// TIA Portal project "Lagerregal_6" (V20)

(* hardware
DEVICE "S7-1500/ET200MP-Station_1"  S7-1500 station
   slot 0: "Profilschiene_0"  Rack  6ES7 590-1***0-0AA0
   slot 1: "PLC_1"  CPU 1513-1 PN  6ES7 513-1AM03-0AB0  V4.0
      slot 3: "CPU-Display_1"  6ES7591-1AA00-0AA0
      slot 32768: "PROFINET-Schnittstelle_1"  X1
         slot 32769: "Port_1"  X1 P1
         slot 32770: "Port_2"  X1 P2
      slot 34817: "Virtual CP interface port_1"  Virtual CP interface port  Virtual CP interface port FW V4.0
   slot 2: "DI 16x24VDC BA_1"  DI 16x24VDC BA  6ES7 521-1BH10-0AA0  V1.1
   slot 3: "DQ 16x24VDC/0.5A ST_1"  DQ 16x24VDC/0.5A ST  6ES7 522-1BH00-0AB0  V2.0
   slot 4: "AI 8xU/I/R/RTD BA_2"  AI 8xU/I/R/RTD BA  6ES7 531-7QF00-0AB0  V1.0
   slot 5: "AI 8xU/I/R/RTD BA_1"  AI 8xU/I/R/RTD BA  6ES7 531-7QF00-0AB0  V1.0
DEVICE "HMI_1"  TP700 Comfort
   slot 0: "HMI_1"  TP700 Comfort  6AV2 124-0GC01-0AX0  17.0.0.0
   slot 1: "HMI_RT_1"  TP700 Comfort  6AV2 124-0GC01-0AX0  17.0.0.0
   slot 5: "HMI_1.IE_CP_1"  PROFINET Interface  17.0.0.0
      slot 1: "PROFINET Schnittstelle_1"  PROFINET Interface
         slot 1: "Port_1"  Port
         slot 2: "Port_2"  Port
   slot 7: "HMI_1.MPI/DP_CP_1"  MPI/DP Interface  17.0.0.0
*)

// ===== PLC "PLC_1"  CPU 1513-1 PN =====

VAR_GLOBAL   // PLC tag table "Standard-Variablentabelle"
   "Clock_Byte" AT %MB0 : Byte;
   "Clock_10Hz" AT %M0.0 : Bool;
   "Clock_5Hz" AT %M0.1 : Bool;
   "Clock_2.5Hz" AT %M0.2 : Bool;
   "Clock_2Hz" AT %M0.3 : Bool;
   "Clock_1.25Hz" AT %M0.4 : Bool;
   "Clock_1Hz" AT %M0.5 : Bool;
   "Clock_0.625Hz" AT %M0.6 : Bool;
   "Clock_0.5Hz" AT %M0.7 : Bool;
END_VAR

VAR_GLOBAL CONSTANT   // PLC tag table "Standard-Variablentabelle"
   "Fachhoehe" : Int := 4800;
   "Fachbreite" : Int := 2962;
   "Offset-Z" : Int := 1800;
   "Offset-X" : Int := 3952;
   "Faecher_pro_Zeile" : Int := 9;
   "Faecher_pro_Spalte" : Int := 6;
   "Anheben_Absenken" : Int := 1000;
END_VAR

VAR_GLOBAL   // PLC tag table "Eingaenge"
   "S1" AT %I0.0 : Bool;   // Not-Aus
   "S2" AT %I0.1 : Bool;   // Anlage ein
   "S3" AT %I0.2 : Bool;   // Starttaster
   "1B1" AT %I0.3 : Bool;   // Sensor 1. Einlassband Anfang
   "1B2" AT %I0.4 : Bool;   // Sensor 1. Einlassband Ende
   "2B1" AT %I0.5 : Bool;   // Sensor 2. Einlassband Anfang
   "2B2" AT %I0.6 : Bool;   // Sensor 2. Einlassband Ende
   "3B1" AT %I0.7 : Bool;   // Sensor 3. Einlassband
   "4B1" AT %I1.0 : Bool;   // Sensor 1. Auslassband
   "5B1" AT %I1.1 : Bool;   // Sensor 2. Auslassband
   "6B1" AT %I1.2 : Bool;   // Endlage Gabel-Kran 1 (links)
   "6B2" AT %I1.3 : Bool;   // Endlage Gabel-Kran 1 (rechts)
   "6B3" AT %I1.4 : Bool;   // Endlage Gabel-Kran 1 (mitte)
   "7B1" AT %I1.5 : Bool;   // Endlage Gabel-Kran 2 (links)
   "7B2" AT %I1.6 : Bool;   // Endlage Gabel-Kran 2 (rechts)
   "7B3" AT %I1.7 : Bool;   // Endlage Gabel-Kran 2 (mitte)
   "2B3" AT %EW30 : Int;   // Kamera am Einlass (Bauteilerkennung)
   "6B4" AT %EW32 : Int;   // X-Achse Kran 1 Ist-Pos
   "6B5" AT %EW34 : Int;   // Z-Achse Kran 1 Ist-Pos
   "7B4" AT %EW36 : Int;   // X-Achse Kran 2 Ist-Pos
   "7B5" AT %EW38 : Int;   // Z-Achse Kran 2 Ist-Pos
END_VAR

VAR_GLOBAL   // PLC tag table "Ausgaenge"
   "H3" AT %Q0.2 : Bool;   // Starttasterleuchte
   "1M1" AT %Q0.3 : Bool;   // 1. Einlassband
   "2M1" AT %Q0.5 : Bool;   // 2. Einlassband
   "3M1" AT %Q0.7 : Bool;   // 3. Einlassband
   "4M1" AT %Q1.0 : Bool;   // 1. Auslassband
   "5M1" AT %Q1.1 : Bool;   // 2. Auslassband
   "6M1" AT %Q1.2 : Bool;   // Gabel-Kran 1 (links)
   "6M2" AT %Q1.3 : Bool;   // Gabel-Kran 1 (rechts)
   "7M1" AT %Q1.5 : Bool;   // Gabel-Kran 2 (links)
   "7M2" AT %Q1.6 : Bool;   // Gabel-Kran 2 (rechts)
   "6M4" AT %AW32 : Int;   // X-Achse Kran 1 Soll-Pos
   "6M5" AT %AW34 : Int;   // Z-Achse Kran 1 Soll-Pos
   "7M4" AT %AW36 : Int;   // X-Achse Kran 2 Soll-Pos
   "7M5" AT %AW38 : Int;   // Z-Achse Kran 2 Soll-Pos
END_VAR

TYPE "typKran_Pos"
   STRUCT
      "X-Ist" : Int;   // X-Achse Kran Ist-Pos
      "X-Soll" : Int;   // X-Achse Kran Soll-Pos
      "X-Rechnen" : Int;   // Zwischenvariable um neue X-Achsen Soll-Pos zu bestimmen
      "X-Skaliert" : Real;
      "Z-Ist" : Int;   // Z-Achse Kran Ist-Pos
      "Z-Soll" : Int;   // Z-Achse Kran Soll-Pos
      "Z-Rechnen" : Int;   // Zwischenvariable um neue Z-Achsen Soll-Pos zu bestimmen
      "Z-Skaliert" : Real;
   END_STRUCT;
END_TYPE

TYPE "typLagerplatz"
   STRUCT
      Flags : Struct
         Belegt : Bool;
         In_Benutzung : Bool;
      END_STRUCT;
      Artikel_Nr : Int;
      Bauteil : Int;
      Zeitstempel : DTL;
      MHD : Date;
   END_STRUCT;
END_TYPE

TYPE "typSchritte"
   STRUCT
      Schritt_Init : Bool;
      Kran : Struct
         Schritt_1 : Bool;
         Schritt_2 : Bool;
         Schritt_3 : Bool;
         Schritt_4 : Bool;
         Schritt_5 : Bool;
      END_STRUCT;
      Kran_Beladen : Struct
         Schritt_1 : Bool;
         Schritt_2 : Bool;
         Schritt_3 : Bool;
         Schritt_4 : Bool;
      END_STRUCT;
      Kran_Entladen : Struct
         Schritt_1 : Bool;
         Schritt_2 : Bool;
         Schritt_3 : Bool;
         Schritt_4 : Bool;
      END_STRUCT;
   END_STRUCT;
END_TYPE

DATA_BLOCK "HMI_Schnittstelle"   // DB100
{ S7_Optimized_Access := 'TRUE' }
VERSION : 0.1
   VAR
      Eingaenge : Struct
         S1 : Bool;   // Not-Aus
         S2 : Bool;   // Anlage ein
         S3 : Bool;   // Starttaster
         "1B1" : Bool;   // Sensor 1. Einlassband Anfang
         "1B2" : Bool;   // Sensor 1. Einlassband Ende
         "2B1" : Bool;   // Sensor 2. Einlassband Anfang
         "2B2" : Bool;   // Sensor 2. Einlassband Ende
         "2B3" : Int;
         "3B1" : Bool;   // Sensor 3. Einlassband
         "4B1" : Bool;   // Sensor 1. Auslassband
         "5B1" : Bool;   // Sensor 2. Auslassband
         "6B1" : Bool;   // Endlage Gabel-Kran 1 (links)
         "6B2" : Bool;   // Endlage Gabel-Kran 1 (rechts)
         "6B3" : Bool;   // Endlage Gabel-Kran 1 (mitte)
         "7B1" : Bool;   // Endlage Gabel-Kran 2 (links)
         "7B2" : Bool;   // Endlage Gabel-Kran 2 (rechts)
         "7B3" : Bool;   // Endlage Gabel-Kran 2 (mitte)
      END_STRUCT;
      Ausgaenge : Struct
         H1 : Bool;   // Starttasterleuchte
         "1M1" : Bool;   // 1. Einlassband
         "2M1" : Bool;   // 2. Einlassband
         "3M1" : Bool;   // 3. Einlassband
         "4M1" : Bool;   // 1. Auslassband
         "5M1" : Bool;   // 2. Auslassband
         "6M1" : Bool;   // Gabel-Kran 1 (links)
         "6M2" : Bool;   // Gabel-Kran 1 (rechts)
         "7M1" : Bool;   // Gabel-Kran 2 (links)
         "7M2" : Bool;   // Gabel-Kran 2 (rechts)
      END_STRUCT;
      Betriebsart : Struct
         Hand : Bool;
         Automatik : Bool;
         Stopp : Bool;
         Einrichten : Bool;
      END_STRUCT;
      Anlagendaten : Struct
         Schrittnummer : UInt;
         Fach_ansteuern : Bool;
         Fach : Int := 1;
         Bauteil : Int;
         Regalplatz_frei : Bool;
         Band_ein : Array[1..3] of Int;
         Band_aus : Array[1..2] of Int;
      END_STRUCT;
      Kraene : Struct
         Kran_1 : Struct
            Kran_Pos : "typKran_Pos";
            Kran_Schritt_Nr : Int;
            Schritt_Beladen : Int;
            Schritt_Entladen : Int;
            Grundstellung : Bool;
            Heimposition : Bool;
            Steht : Bool;
            Beladen : Bool;
         END_STRUCT;
         Kran_2 : Struct
            Kran_Pos : "typKran_Pos";
            Kran_Schritt_Nr : Int;
            Schritt_Beladen : Int;
            Schritt_Entladen : Int;
            Grundstellung : Bool;
            Heimposition : Bool;
            Steht : Bool;
            Beladen : Bool;
         END_STRUCT;
      END_STRUCT;
      HMI : Struct
         "X-Pos" : Bool;   // X-Achse-Inkrement erhöhen Schalter
         "X-Neg" : Bool;   // X-Achse-Inkrement verringern Schalter
         "Z-Pos" : Bool;   // Z-Achse-Inkrement erhöhen Schalter
         "Z-Neg" : Bool;   // Z-Achse-Inkrement verringern Schalter
         Inkrement : UInt;   // Inkrement Schrittgröße für Achsen
      END_STRUCT;
      Bitmeldungen : Word;
   END_VAR
BEGIN
   // Kraene.Kran_1.Kran_Pos."X-Ist" : X-Achse Kran 1 Ist-Pos
   // Kraene.Kran_1.Kran_Pos."Z-Ist" : Z-Achse Kran 1 Ist-Pos
   // Kraene.Kran_2.Kran_Pos."X-Ist" : X-Achse Kran 2 Ist-Pos
   // Kraene.Kran_2.Kran_Pos."Z-Ist" : Z-Achse Kran 2 Ist-Pos
   // Kraene.Kran_1.Kran_Pos."X-Soll" : X-Achse Kran 1 Soll-Pos
   // Kraene.Kran_1.Kran_Pos."Z-Soll" : Z-Achse Kran 1 Soll-Pos
   // Kraene.Kran_2.Kran_Pos."X-Soll" : X-Achse Kran 2 Soll-Pos
   // Kraene.Kran_2.Kran_Pos."Z-Soll" : Z-Achse Kran 2 Soll-Pos
END_DATA_BLOCK

DATA_BLOCK "Warenlager"   // DB101
{ S7_Optimized_Access := 'TRUE' }
VERSION : 0.1
   VAR
      Lager : Array[0..54] of "typLagerplatz";
   END_VAR
BEGIN
END_DATA_BLOCK

// folder: Anlagedaten

DATA_BLOCK "IDB_Anlage"   // DB1
{ S7_Optimized_Access := 'TRUE' }
VERSION : 0.1
// stored: InstanceOfName Ein_Anlage
"Ein_Anlage"
BEGIN
END_DATA_BLOCK

// folder: Bandsteuerung

DATA_BLOCK "IDB_Baender"   // DB20
{ S7_Optimized_Access := 'TRUE' }
VERSION : 0.1
// stored: InstanceOfName Ein_Baender
"Ein_Baender"
BEGIN
END_DATA_BLOCK

DATA_BLOCK "IDB_Bandsteuerung"   // DB21
{ S7_Optimized_Access := 'TRUE' }
VERSION : 0.1
// stored: InstanceOfName Bandsteuerung
"Bandsteuerung"
BEGIN
END_DATA_BLOCK

// folder: HMI

DATA_BLOCK "IDB_Einrichtbetrieb"   // DB3
{ S7_Optimized_Access := 'TRUE' }
VERSION : 0.1
// stored: InstanceOfName Prog_Einrichtbetrieb
"Prog_Einrichtbetrieb"
BEGIN
END_DATA_BLOCK

DATA_BLOCK "IDB_HMI"   // DB10
{ S7_Optimized_Access := 'TRUE' }
VERSION : 0.1
// stored: InstanceOfName Ein_HMI
"Ein_HMI"
BEGIN
END_DATA_BLOCK

// folder: Kransteuerung

DATA_BLOCK "IDB_Kran_beladen"   // DB25
{ S7_Optimized_Access := 'TRUE' }
VERSION : 0.1
// stored: InstanceOfName FC_Kran_beladen
"FC_Kran_beladen"
BEGIN
END_DATA_BLOCK

DATA_BLOCK "IDB_Kran"   // DB30
{ S7_Optimized_Access := 'TRUE' }
VERSION : 0.1
// stored: InstanceOfName Ein_Kran
"Ein_Kran"
BEGIN
END_DATA_BLOCK

DATA_BLOCK "IDB_Automatik_einlagern"   // DB50
{ S7_Optimized_Access := 'TRUE' }
VERSION : 0.1
// stored: InstanceOfName Prog_Automatik_einlagern
"Prog_Automatik_einlagern"
BEGIN
END_DATA_BLOCK

DATA_BLOCK "IDB_Automatik_auslagern"   // DB60
{ S7_Optimized_Access := 'TRUE' }
VERSION : 0.1
// stored: InstanceOfName Prog_Automatik_auslagern
"Prog_Automatik_auslagern"
BEGIN
END_DATA_BLOCK

// folder: (top level)

FUNCTION_BLOCK "Prog_Schrittkette"   // FB1234, FBD
{ S7_Optimized_Access := 'TRUE' }
VERSION : 0.1
   VAR_INPUT
      eAutomatik : Bool;   // Automatikmodus
      eAusschalten : Bool;   // Ausschalten der Schrittkette
      T_1_2 : Bool;
      T_2_3 : Bool;
      T_3_4 : Bool := TRUE;
      T_4_5 : Bool := TRUE;
      T_5_6 : Bool := TRUE;
      T_6_7 : Bool := TRUE;
      T_7_8 : Bool := TRUE;
      T_8_9 : Bool := TRUE;
      T_9_10 : Bool := TRUE;
      T_10_1 : Bool := TRUE;
   END_VAR
   VAR_OUTPUT
      aSchrittnummer : Int;
   END_VAR
   VAR
      Step_1 : Bool;
      Step_2 : Bool;
      Step_3 : Bool;
      Step_4 : Bool;
      Step_5 : Bool;
      Step_6 : Bool;
      Step_7 : Bool;
      Step_8 : Bool;
      Step_9 : Bool;
      Step_10 : Bool;
   END_VAR
BEGIN

REGION Network 1: Step 1
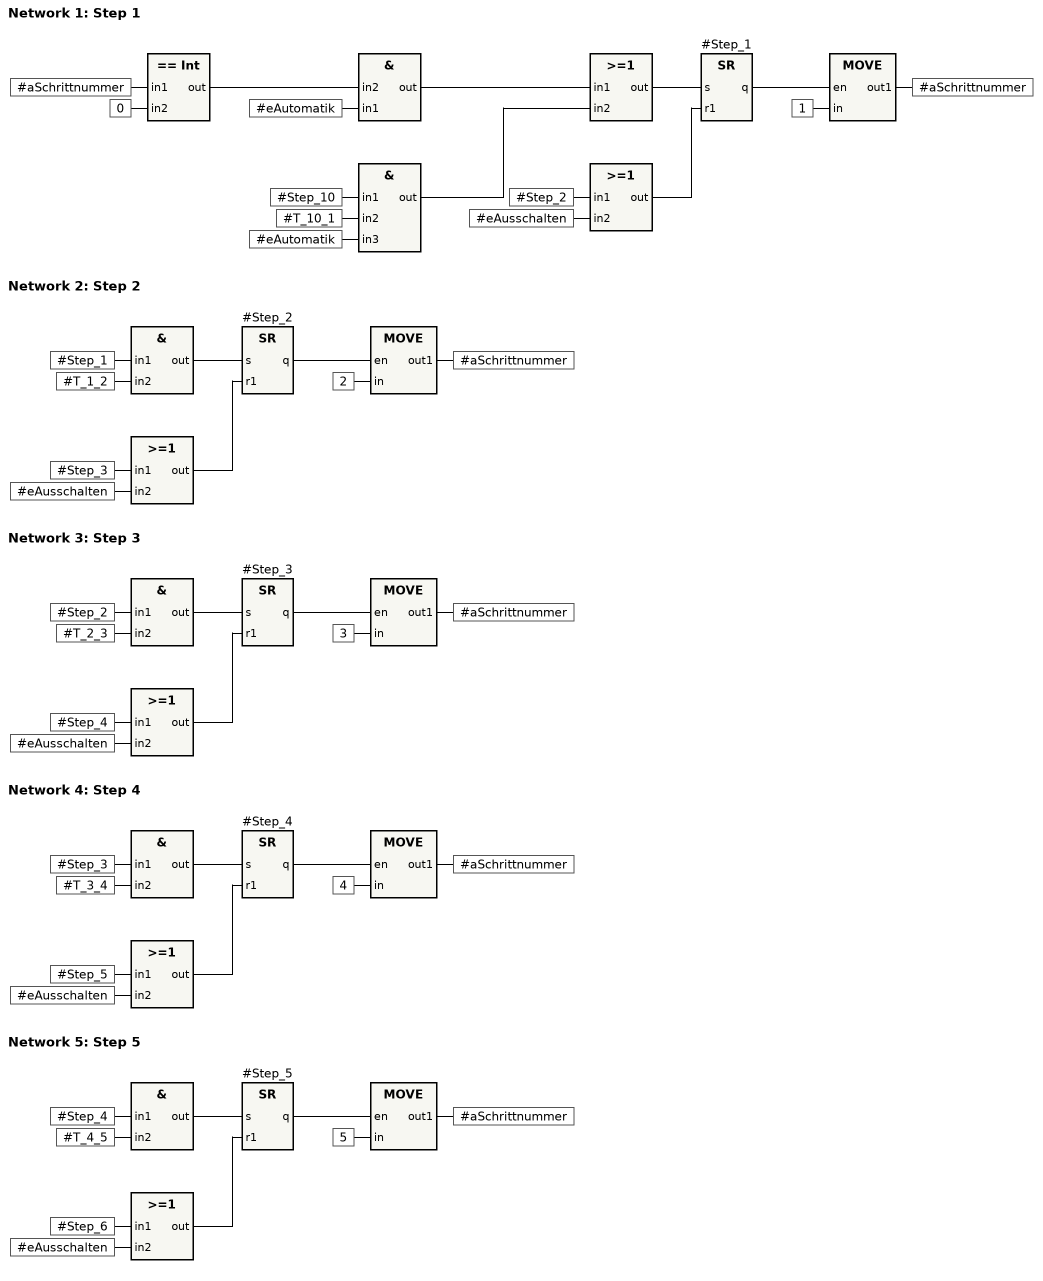
   IF ((#aSchrittnummer = 0) AND #eAutomatik) OR (#Step_10 AND #T_10_1 AND #eAutomatik) THEN
       #Step_1 := TRUE;   // SR flip-flop
   END_IF;
   IF #Step_2 OR #eAusschalten THEN #Step_1 := FALSE; END_IF;
   IF #Step_1 THEN #aSchrittnummer := 1; END_IF;
END_REGION

REGION Network 2: Step 2
   IF #Step_1 AND #T_1_2 THEN
       #Step_2 := TRUE;   // SR flip-flop
   END_IF;
   IF #Step_3 OR #eAusschalten THEN #Step_2 := FALSE; END_IF;
   IF #Step_2 THEN #aSchrittnummer := 2; END_IF;
END_REGION

REGION Network 3: Step 3
   IF #Step_2 AND #T_2_3 THEN
       #Step_3 := TRUE;   // SR flip-flop
   END_IF;
   IF #Step_4 OR #eAusschalten THEN #Step_3 := FALSE; END_IF;
   IF #Step_3 THEN #aSchrittnummer := 3; END_IF;
END_REGION

REGION Network 4: Step 4
   IF #Step_3 AND #T_3_4 THEN
       #Step_4 := TRUE;   // SR flip-flop
   END_IF;
   IF #Step_5 OR #eAusschalten THEN #Step_4 := FALSE; END_IF;
   IF #Step_4 THEN #aSchrittnummer := 4; END_IF;
END_REGION

REGION Network 5: Step 5
   IF #Step_4 AND #T_4_5 THEN
       #Step_5 := TRUE;   // SR flip-flop
   END_IF;
   IF #Step_6 OR #eAusschalten THEN #Step_5 := FALSE; END_IF;
   IF #Step_5 THEN #aSchrittnummer := 5; END_IF;
END_REGION

REGION Network 6: Step 6
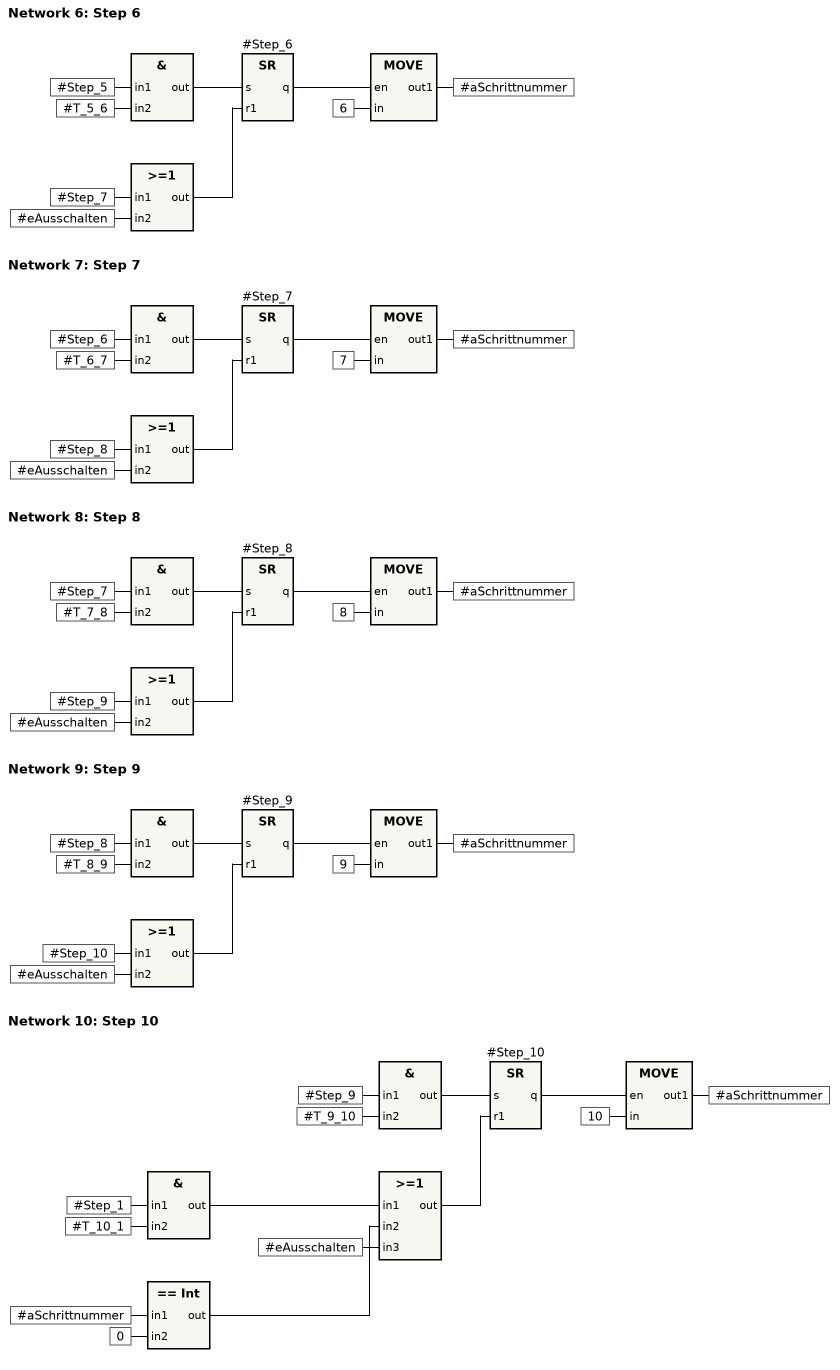
   IF #Step_5 AND #T_5_6 THEN
       #Step_6 := TRUE;   // SR flip-flop
   END_IF;
   IF #Step_7 OR #eAusschalten THEN #Step_6 := FALSE; END_IF;
   IF #Step_6 THEN #aSchrittnummer := 6; END_IF;
END_REGION

REGION Network 7: Step 7
   IF #Step_6 AND #T_6_7 THEN
       #Step_7 := TRUE;   // SR flip-flop
   END_IF;
   IF #Step_8 OR #eAusschalten THEN #Step_7 := FALSE; END_IF;
   IF #Step_7 THEN #aSchrittnummer := 7; END_IF;
END_REGION

REGION Network 8: Step 8
   IF #Step_7 AND #T_7_8 THEN
       #Step_8 := TRUE;   // SR flip-flop
   END_IF;
   IF #Step_9 OR #eAusschalten THEN #Step_8 := FALSE; END_IF;
   IF #Step_8 THEN #aSchrittnummer := 8; END_IF;
END_REGION

REGION Network 9: Step 9
   IF #Step_8 AND #T_8_9 THEN
       #Step_9 := TRUE;   // SR flip-flop
   END_IF;
   IF #Step_10 OR #eAusschalten THEN #Step_9 := FALSE; END_IF;
   IF #Step_9 THEN #aSchrittnummer := 9; END_IF;
END_REGION

REGION Network 10: Step 10
   IF #Step_9 AND #T_9_10 THEN
       #Step_10 := TRUE;   // SR flip-flop
   END_IF;
   IF (#Step_1 AND #T_10_1) OR (#aSchrittnummer = 0) OR #eAusschalten THEN #Step_10 := FALSE; END_IF;
   IF #Step_10 THEN #aSchrittnummer := 10; END_IF;
END_REGION

REGION Network 11: Schrittkette beenden, wenn der Automatikmodus beendet wird
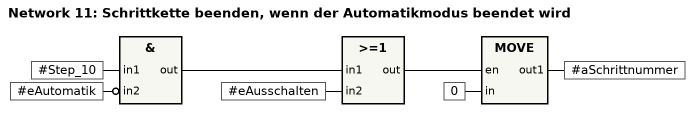
   IF (#Step_10 AND NOT #eAutomatik) OR #eAusschalten THEN #aSchrittnummer := 0; END_IF;
END_REGION
END_FUNCTION_BLOCK

FUNCTION "Analog_Test" : Void   // FC2, FBD
{ S7_Optimized_Access := 'TRUE' }
VERSION : 0.1
   VAR_INPUT
      X_skaliert : Real;
      Z_skaliert : Real;
   END_VAR
   VAR_OUTPUT
      Soll_X : Int;
      Soll_Z : Int;
   END_VAR
   VAR_TEMP
      normierter_Wert_X : Real;
      normierter_Wert_Z : Real;
   END_VAR
BEGIN

REGION Network 1
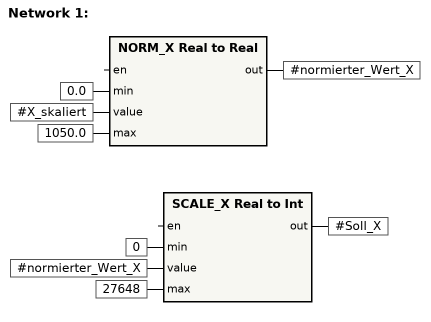
   #normierter_Wert_X := NORM_X(MIN := 0.0, VALUE := #X_skaliert, MAX := 1050.0);
   #Soll_X := SCALE_X(MIN := 0, VALUE := #normierter_Wert_X, MAX := 27648);
END_REGION

REGION Network 2 (SCL)
   #normierter_Wert_Z := NORM_X(MIN := 0.0, VALUE := #Z_skaliert, MAX := 662.5);
   #Soll_Z := SCALE_X(MIN := 0, VALUE := #normierter_Wert_Z, MAX := 27648);
END_REGION
END_FUNCTION

FUNCTION "Generiere_Zufallszahl" : UDInt   // FC3, SCL
{ S7_Optimized_Access := 'TRUE' }
VERSION : 0.1
   VAR_INPUT
      iObergrenze : UDInt;
      iUntergrenze : UDInt;
   END_VAR
   VAR_OUTPUT
      aFehler : Int;   // Rückgabewert von RD_LOC_T, falls es einen Fehler gab beim erzeugen der Zufallszahl.
   END_VAR
   VAR_TEMP
      tmpZeitstempel : DTL;
      tmpZeit_als_Zahl : UDInt;   // Nanosekunde aus dem Zeitstempel.
   END_VAR
   // Ret_Val : Eine Zufallszahl zwischen der oberen und unteren Grenze.
BEGIN
   (*
       Die zu erzeugende Zufallszahl
   *)
   IF
       // #iObergrenze >= 999 OR
       #iUntergrenze >= #iObergrenze OR
       // Die Obergrenze minus der Untergrenze muss mindestens 2 ergeben.
       (#iObergrenze - #iUntergrenze) <= 1
   THEN
       #aFehler := 2;
       #Generiere_Zufallszahl := 0;
       RETURN;
   END_IF;


   #aFehler := RD_LOC_T(#tmpZeitstempel);
   #tmpZeit_als_Zahl := (#tmpZeitstempel.HOUR * 10000000) + (#tmpZeitstempel.MINUTE * 100000) + (#tmpZeitstempel.SECOND * 1000) + #tmpZeitstempel.NANOSECOND;


   // Hier wird die zu erzeugende 'Zufallszahl' zurückgegeben.
   #Generiere_Zufallszahl := (#tmpZeit_als_Zahl MOD (#iObergrenze - #iUntergrenze)) + #iUntergrenze;
END_FUNCTION

FUNCTION "Analogwerte" : Void   // FC25, FBD
{ S7_Optimized_Access := 'TRUE' }
VERSION : 0.1
   VAR_INPUT
      Ist_X : Int;
      Ist_Z : Int;
   END_VAR
   VAR_OUTPUT
      X_skaliert : Real;
      Z_skaliert : Real;
   END_VAR
   VAR_TEMP
      normierter_Wert_X : Real;
      normierter_Wert_Z : Real;
   END_VAR
BEGIN

REGION Network 1: Stapler Umwandlung X-Achse in cm
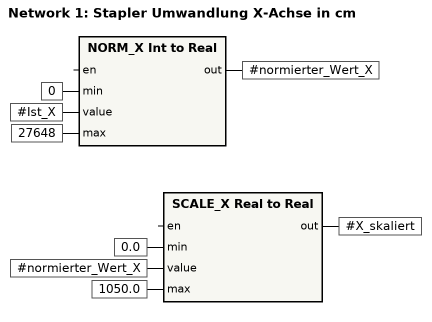
   #normierter_Wert_X := NORM_X(MIN := 0, VALUE := #Ist_X, MAX := 27648);
   #X_skaliert := SCALE_X(MIN := 0.0, VALUE := #normierter_Wert_X, MAX := 1050.0);
END_REGION

REGION Network 2 (SCL): Stapler Umwandlung Z-Achse in cm
   #normierter_Wert_Z := NORM_X(MIN := 0, VALUE := #Ist_Z, MAX := 27648);
   #Z_skaliert := SCALE_X(MIN := 0.0, VALUE := #normierter_Wert_Z, MAX := 662.5);
END_REGION
END_FUNCTION

FUNCTION "Berechne_Offset" : Void   // FC5000, SCL
{ S7_Optimized_Access := 'TRUE' }
VERSION : 0.1
   VAR_INPUT
      eFach_Nr : DInt;
      eFach_Anzahl : DInt;
      eFach_Breite : DInt;
      eFach_Hoehe : DInt;
      eOffset_X : DInt;
      eOffset_Z : DInt;
   END_VAR
   VAR_OUTPUT
      aPos_X : DInt;
      aPos_Z : DInt;
   END_VAR
BEGIN
   (*
      Der Baustein berechnet die Koordinaten (X,Z) eines Fachs
      in Abhängigkeit von einer Fachnummer

      Der Baustein ist universell einsetzbar für alle gleichhbleibenden Raster.
   *)

   // Position setzen
   IF #eFach_Nr > 0 THEN
       #aPos_X := ((#eFach_Nr - 1) MOD #eFach_Anzahl) * #eFach_Breite + #eOffset_X;
       #aPos_Z := ((#eFach_Nr - 1) / #eFach_Anzahl) * #eFach_Hoehe + #eOffset_Z;
   ELSE
       #aPos_X := #aPos_Z := 0;
   END_IF;
END_FUNCTION

ORGANIZATION_BLOCK "Main"   // OB1, FBD, ProgramCycle
TITLE = "Main Program Sweep (Cycle)"
{ S7_Optimized_Access := 'TRUE' }
VERSION : 0.1
   VAR_INPUT
      Initial_Call : Bool;   // Initial call of this OB
      Remanence : Bool;   // =True, if remanent data are available
   END_VAR
BEGIN

REGION Network 1: Eingang von Anlagesensorik
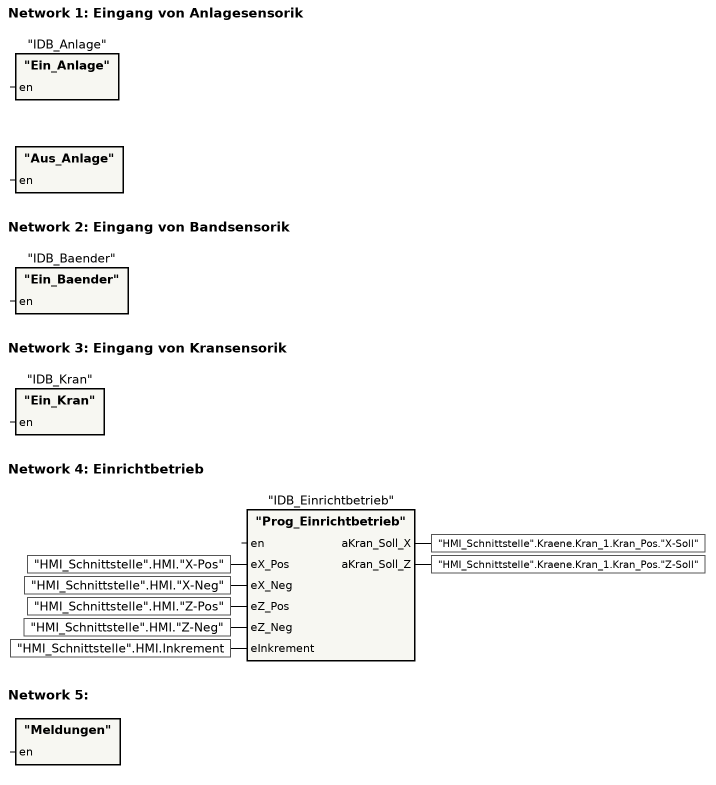
   "IDB_Anlage"();   // "Ein_Anlage"
   "Aus_Anlage"();
END_REGION

REGION Network 2: Eingang von Bandsensorik
   "IDB_Baender"();   // "Ein_Baender"
END_REGION

REGION Network 3: Eingang von Kransensorik
   "IDB_Kran"();   // "Ein_Kran"
END_REGION

REGION Network 4: Einrichtbetrieb
   "IDB_Einrichtbetrieb"(eX_Pos := "HMI_Schnittstelle".HMI."X-Pos",   // "Prog_Einrichtbetrieb"
                         eX_Neg := "HMI_Schnittstelle".HMI."X-Neg",
                         eZ_Pos := "HMI_Schnittstelle".HMI."Z-Pos",
                         eZ_Neg := "HMI_Schnittstelle".HMI."Z-Neg",
                         eInkrement := "HMI_Schnittstelle".HMI.Inkrement,
                         aKran_Soll_X => "HMI_Schnittstelle".Kraene.Kran_1.Kran_Pos."X-Soll",
                         aKran_Soll_Z => "HMI_Schnittstelle".Kraene.Kran_1.Kran_Pos."Z-Soll");
END_REGION

REGION Network 5
   "Meldungen"();
END_REGION
END_ORGANIZATION_BLOCK

// folder: Anlagedaten

FUNCTION_BLOCK "Ein_Anlage"   // FB1, FBD
{ S7_Optimized_Access := 'TRUE' }
VERSION : 0.1
BEGIN

REGION Network 1: Schalter einlesen
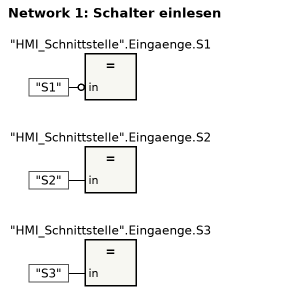
   "HMI_Schnittstelle".Eingaenge.S1 := NOT "S1";
   "HMI_Schnittstelle".Eingaenge.S2 := "S2";
   "HMI_Schnittstelle".Eingaenge.S3 := "S3";
END_REGION
END_FUNCTION_BLOCK

FUNCTION "Aus_Anlage" : Void   // FC1, FBD
{ S7_Optimized_Access := 'TRUE' }
VERSION : 0.1
BEGIN

REGION Network 1 (SCL): Leuchte Starttaster
   "HMI_Schnittstelle".Ausgaenge.H1 := "HMI_Schnittstelle".Eingaenge.S2;
END_REGION
END_FUNCTION

// folder: Bandsteuerung

FUNCTION_BLOCK "Ein_Baender"   // FB20, FBD
{ S7_Optimized_Access := 'TRUE' }
VERSION : 0.1
BEGIN

REGION Network 1 (SCL): Sensoren Einlass
   "HMI_Schnittstelle".Eingaenge."1B1" := NOT "1B1";
   "HMI_Schnittstelle".Eingaenge."1B2" := NOT "1B2";
   "HMI_Schnittstelle".Eingaenge."2B1" := NOT "2B1";
   "HMI_Schnittstelle".Eingaenge."2B2" := NOT "2B2";
   "HMI_Schnittstelle".Eingaenge."2B3" := "2B3";
   "HMI_Schnittstelle".Eingaenge."3B1" := NOT "3B1";
END_REGION

REGION Network 2 (SCL): Sensoren Auslass
   "HMI_Schnittstelle".Eingaenge."4B1" := NOT "4B1";
   "HMI_Schnittstelle".Eingaenge."5B1" := NOT "5B1";
END_REGION
END_FUNCTION_BLOCK

FUNCTION_BLOCK "Bandsteuerung"   // FB21, FBD
{ S7_Optimized_Access := 'TRUE' }
VERSION : 0.1
   VAR
      FTRIG_MDB_1B1 : F_TRIG;
      FTRIG_MDB_1B2 : F_TRIG;
      FTRIG_MDB_2B1 : F_TRIG;
      FTRIG_MDB_2B2 : F_TRIG;
      FTRIG_MDB_5B1 : F_TRIG;
      RTRIG_MDB_5B1 : R_TRIG;
      Band_belegt : Bool;
   END_VAR
BEGIN

REGION Network 1 (SCL): Flankenabfragen
   #FTRIG_MDB_1B1(CLK := "HMI_Schnittstelle".Eingaenge."1B1");
   #FTRIG_MDB_1B2(CLK:="HMI_Schnittstelle".Eingaenge."1B2");
   #FTRIG_MDB_2B1(CLK := "HMI_Schnittstelle".Eingaenge."2B1");
   #FTRIG_MDB_2B2(CLK := "HMI_Schnittstelle".Eingaenge."2B2");
   #FTRIG_MDB_5B1(CLK := "HMI_Schnittstelle".Eingaenge."5B1");
   #RTRIG_MDB_5B1(CLK := "HMI_Schnittstelle".Eingaenge."5B1");
END_REGION

REGION Network 2: Einlasssteuerung (Band 1)
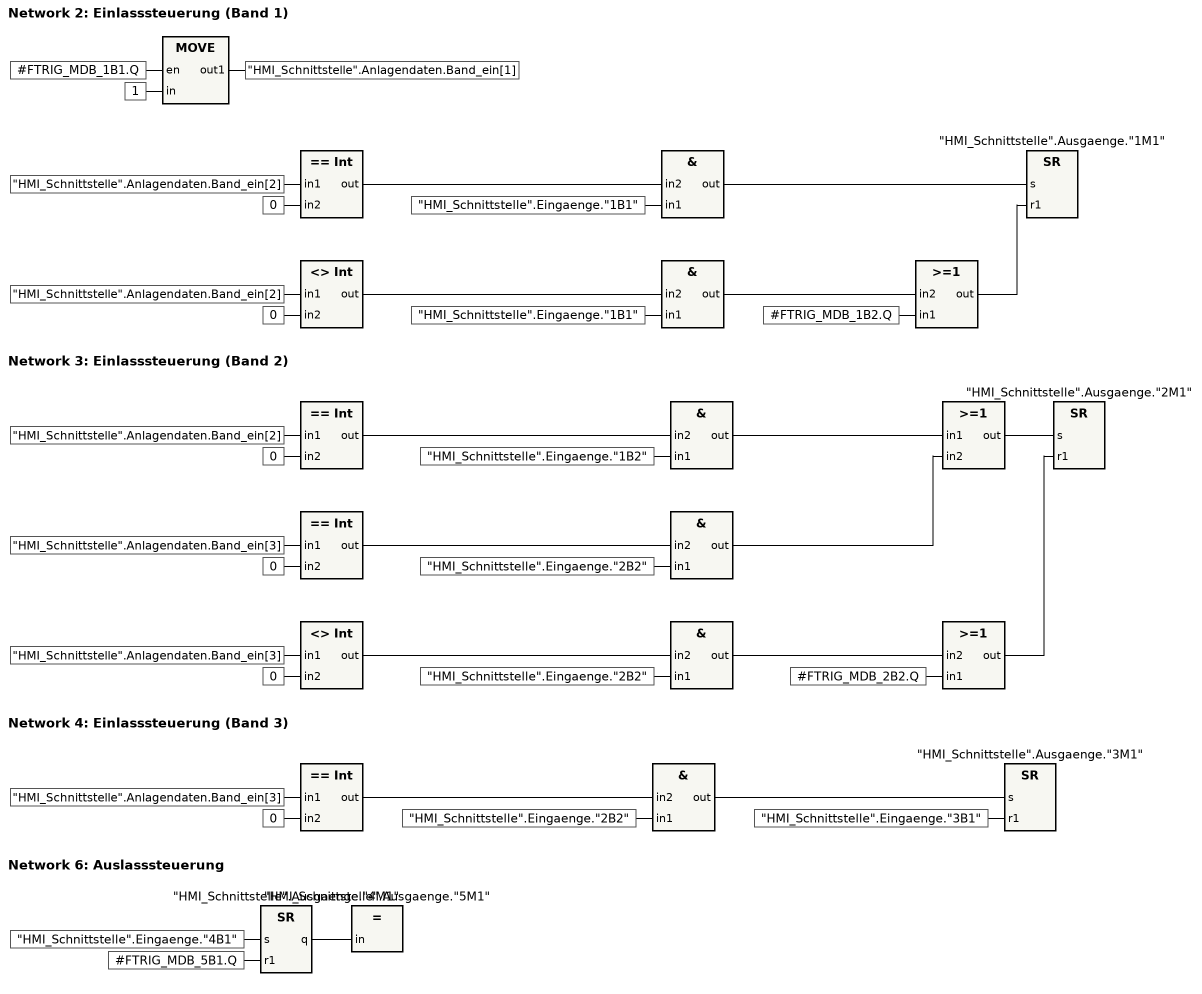
   IF #FTRIG_MDB_1B1.Q THEN "HMI_Schnittstelle".Anlagendaten.Band_ein[1] := 1; END_IF;
   IF ("HMI_Schnittstelle".Anlagendaten.Band_ein[2] = 0) AND "HMI_Schnittstelle".Eingaenge."1B1" THEN
       "HMI_Schnittstelle".Ausgaenge."1M1" := TRUE;   // SR flip-flop
   END_IF;
   IF (("HMI_Schnittstelle".Anlagendaten.Band_ein[2] <> 0) AND "HMI_Schnittstelle".Eingaenge."1B1") OR #FTRIG_MDB_1B2.Q THEN
       "HMI_Schnittstelle".Ausgaenge."1M1" := FALSE;
   END_IF;
END_REGION

REGION Network 3: Einlasssteuerung (Band 2)
   IF (("HMI_Schnittstelle".Anlagendaten.Band_ein[2] = 0) AND "HMI_Schnittstelle".Eingaenge."1B2") OR (("HMI_Schnittstelle".Anlagendaten.Band_ein[3] = 0) AND "HMI_Schnittstelle".Eingaenge."2B2") THEN
       "HMI_Schnittstelle".Ausgaenge."2M1" := TRUE;   // SR flip-flop
   END_IF;
   IF (("HMI_Schnittstelle".Anlagendaten.Band_ein[3] <> 0) AND "HMI_Schnittstelle".Eingaenge."2B2") OR #FTRIG_MDB_2B2.Q THEN
       "HMI_Schnittstelle".Ausgaenge."2M1" := FALSE;
   END_IF;
END_REGION

REGION Network 4: Einlasssteuerung (Band 3)
   IF ("HMI_Schnittstelle".Anlagendaten.Band_ein[3] = 0) AND "HMI_Schnittstelle".Eingaenge."2B2" THEN
       "HMI_Schnittstelle".Ausgaenge."3M1" := TRUE;   // SR flip-flop
   END_IF;
   IF "HMI_Schnittstelle".Eingaenge."3B1" THEN "HMI_Schnittstelle".Ausgaenge."3M1" := FALSE; END_IF;
END_REGION

REGION Network 5 (SCL): Bandbelegung
   IF #FTRIG_MDB_2B1.Q THEN
       "HMI_Schnittstelle".Anlagendaten.Band_ein[2] := "HMI_Schnittstelle".Anlagendaten.Band_ein[1];
       "HMI_Schnittstelle".Anlagendaten.Band_ein[1] := 0;
   END_IF;

   IF #FTRIG_MDB_2B2.Q THEN
       "HMI_Schnittstelle".Anlagendaten.Band_ein[3] := "HMI_Schnittstelle".Anlagendaten.Band_ein[2];
       "HMI_Schnittstelle".Anlagendaten.Band_ein[2] := 0;
   END_IF;

   IF "HMI_Schnittstelle".Eingaenge."2B3" <> 0 AND "HMI_Schnittstelle".Anlagendaten.Band_ein[2] = 1 THEN
       "HMI_Schnittstelle".Anlagendaten.Band_ein[2] := "HMI_Schnittstelle".Eingaenge."2B3";
   END_IF;
END_REGION

REGION Network 6: Auslasssteuerung
   IF "HMI_Schnittstelle".Eingaenge."4B1" THEN
       "HMI_Schnittstelle".Ausgaenge."4M1" := TRUE;   // SR flip-flop
   END_IF;
   IF #FTRIG_MDB_5B1.Q THEN "HMI_Schnittstelle".Ausgaenge."4M1" := FALSE; END_IF;
   "HMI_Schnittstelle".Ausgaenge."5M1" := "HMI_Schnittstelle".Ausgaenge."4M1";
END_REGION

REGION Network 7 (SCL): Bandbelegung
   IF "HMI_Schnittstelle".Eingaenge."5B1" THEN
       "HMI_Schnittstelle".Anlagendaten.Band_aus[2] := "HMI_Schnittstelle".Anlagendaten.Band_aus[1];
       "HMI_Schnittstelle".Anlagendaten.Band_aus[1] := 0;
   END_IF;

   IF #RTRIG_MDB_5B1.Q THEN
       "HMI_Schnittstelle".Anlagendaten.Band_aus[2] := 0;
   END_IF;
END_REGION
END_FUNCTION_BLOCK

FUNCTION "Aus_Baender" : Void   // FC20, FBD
{ S7_Optimized_Access := 'TRUE' }
VERSION : 0.1
BEGIN

REGION Network 1 (SCL): Bänder Einlass
   "1M1" := "HMI_Schnittstelle".Ausgaenge."1M1";
   "2M1" := "HMI_Schnittstelle".Ausgaenge."2M1";
   "3M1" := "HMI_Schnittstelle".Ausgaenge."3M1";
END_REGION

REGION Network 2 (SCL): Bänder Auslass
   "4M1" := "HMI_Schnittstelle".Ausgaenge."4M1";
   "5M1" := "HMI_Schnittstelle".Ausgaenge."5M1";
END_REGION
END_FUNCTION

ORGANIZATION_BLOCK "Main_Baender"   // OB124, FBD, ProgramCycle
TITLE = "Main Program Sweep (Cycle)"
{ S7_Optimized_Access := 'TRUE' }
VERSION : 0.1
   VAR_INPUT
      Initial_Call : Bool;   // Initial call of this OB
      Remanence : Bool;   // =True, if remanent data are available
   END_VAR
BEGIN

REGION Network 1
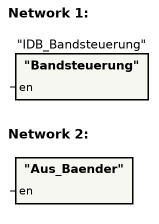
   "IDB_Bandsteuerung"();   // "Bandsteuerung"
END_REGION

REGION Network 2
   "Aus_Baender"();
END_REGION
END_ORGANIZATION_BLOCK

// folder: HMI

FUNCTION_BLOCK "Prog_Einrichtbetrieb"   // FB3, FBD
{ S7_Optimized_Access := 'TRUE' }
VERSION : 0.1
   VAR_INPUT
      eX_Pos : Bool;
      eX_Neg : Bool;
      eZ_Pos : Bool;
      eZ_Neg : Bool;
      eInkrement : UInt;
   END_VAR
   VAR_OUTPUT
      aKran_Soll_X : Int;
      aKran_Soll_Z : Int;
   END_VAR
   VAR
      "PTRIG_MDB_X-Pos" : R_TRIG;
      "PTRIG_MDB_X-Neg" : R_TRIG;
      "PTRIG_MDB_Z-Pos" : R_TRIG;
      "PTRIG_MDB_Z-Neg" : R_TRIG;
   END_VAR
BEGIN

REGION Network 1 (SCL): Button Flanken erfassen
   #"PTRIG_MDB_X-Pos"(CLK := #eX_Pos);
   #"PTRIG_MDB_X-Neg"(CLK := #eX_Neg);

   #"PTRIG_MDB_Z-Pos"(CLK := #eZ_Pos);
   #"PTRIG_MDB_Z-Neg"(CLK := #eZ_Neg);
END_REGION

REGION Network 2 (SCL): Achsen inkrementieren
   // X-Achse Inkrementieren
   IF #"PTRIG_MDB_X-Pos".Q THEN
       #aKran_Soll_X += UINT_TO_INT(#eInkrement);
   END_IF;

   IF #"PTRIG_MDB_X-Neg".Q THEN
       #aKran_Soll_X -= UINT_TO_INT(#eInkrement);
   END_IF;


   // Z-Achse Inkrementieren
   IF #"PTRIG_MDB_Z-Pos".Q THEN
       #aKran_Soll_Z += UINT_TO_INT(#eInkrement);
   END_IF;

   IF #"PTRIG_MDB_Z-Neg".Q THEN
       #aKran_Soll_Z -= UINT_TO_INT(#eInkrement);
   END_IF;
END_REGION
END_FUNCTION_BLOCK

FUNCTION_BLOCK "Ein_HMI"   // FB10, FBD
{ S7_Optimized_Access := 'TRUE' }
VERSION : 0.1
BEGIN
END_FUNCTION_BLOCK

FUNCTION "Meldungen" : Void   // FC10, SCL
{ S7_Optimized_Access := 'TRUE' }
VERSION : 0.1
BEGIN
   // Slice Zugriff programmieren
   // d.h. wir können auf die Einzelbits einer Ganzzahlvariable (INT, DINT, etc.)
   // bzw. einer Bitfolge (Byte, Word, etc.) zugreifen.

   // Bits:        Variable.%X0
   // Bytes:       Variable.%B0
   // Word:        Variable.%W0
   // DWord:       Variable.%D0


   "HMI_Schnittstelle".Bitmeldungen.%X0 := "HMI_Schnittstelle".Eingaenge.S2;
   "HMI_Schnittstelle".Bitmeldungen.%X1 := "HMI_Schnittstelle".Eingaenge.S1;
   "HMI_Schnittstelle".Bitmeldungen.%X2 := "HMI_Schnittstelle".Betriebsart.Hand;
   "HMI_Schnittstelle".Bitmeldungen.%X3 := "HMI_Schnittstelle".Betriebsart.Automatik;
END_FUNCTION

// folder: Kransteuerung

FUNCTION_BLOCK "FC_Kran_beladen"   // FB25, FBD
{ S7_Optimized_Access := 'TRUE' }
VERSION : 0.1
   VAR_INPUT
      eKran_Ist_X : Int;
      eKran_Ist_Z : Int;
      eKran_Soll_X : Int;
      eKran_Soll_Z : Int;
      eGabel_Mitte : Bool;
      eSchrittnummer : UInt;
      ePalette_abholbereit : Bool;
   END_VAR
   VAR_OUTPUT
      aKran_Soll_X : Int;
      aKran_Soll_Z : Int;
      aGabel_Links : Bool;
      aGabel_Rechts : Bool;
      aBeladen : Bool;
   END_VAR
   VAR_TEMP
      tmpRD_T_ERR : Int;
   END_VAR
BEGIN

REGION Network 1 (SCL): Gabel links ausfahren
   #aGabel_Links := #eSchrittnummer = 2 OR #eSchrittnummer = 3;
END_REGION

REGION Network 2 (SCL): Gabel rechts ausfahren
   #aGabel_Rechts := #eSchrittnummer = 6 OR #eSchrittnummer = 7;
END_REGION

REGION Network 3 (SCL): Z-Achse Kran Soll-Pos
   // Einrichtbetrieb
   IF "HMI_Schnittstelle".Betriebsart.Einrichten THEN
       #aKran_Soll_Z := "HMI_Schnittstelle".Kraene.Kran_1.Kran_Pos."Z-Soll";

   // Automatikbetrieb
   ELSIF "HMI_Schnittstelle".Betriebsart.Automatik THEN

       CASE #eSchrittnummer OF
           3:
               // Palette aus Grundstellung anheben
               #aKran_Soll_Z := "Anheben_Absenken" + 2;
           5:
               //Fach mit Nummer anfahren
               #aKran_Soll_Z := #eKran_Soll_Z;
           7:
               // Palette in Regal einlagern
               #aKran_Soll_Z := #eKran_Soll_Z - "Anheben_Absenken";
           9:
               // Stapler in Grundstellung
               #aKran_Soll_Z := 0;
           ELSE:
               ;
       END_CASE;

   END_IF;
END_REGION

REGION Network 4 (SCL): Flag Kran beladen
   IF "HMI_Schnittstelle".Betriebsart.Einrichten THEN
       #aBeladen := FALSE;
   END_IF;


   IF #ePalette_abholbereit
       AND #"eKran_Ist_X" = 0
       AND #"eKran_Ist_Z" >= "Anheben_Absenken"
       AND #eGabel_Mitte
   THEN
       #aBeladen := TRUE;

       "HMI_Schnittstelle".Anlagendaten.Bauteil := "HMI_Schnittstelle".Anlagendaten.Band_ein[3];
       "HMI_Schnittstelle".Anlagendaten.Band_ein[3] := 0;
   END_IF;


   IF #"eKran_Ist_X" = #eKran_Soll_X
       AND #"eKran_Ist_Z" = #eKran_Soll_Z
       AND #eGabel_Mitte
       AND #aBeladen
   THEN
       "Warenlager".Lager["HMI_Schnittstelle".Anlagendaten.Fach].Flags.In_Benutzung := TRUE;
   END_IF;


   IF #"eKran_Ist_X" = #eKran_Soll_X
       AND #"eKran_Ist_Z" = #eKran_Soll_Z - "Anheben_Absenken"
       AND #aBeladen
   THEN
       // Wenn die Palette eingelagert wurde, schreibe die Info über das Bauteil ins Array.
       "Warenlager".Lager["HMI_Schnittstelle".Anlagendaten.Fach].Flags.Belegt := TRUE;
       "Warenlager".Lager["HMI_Schnittstelle".Anlagendaten.Fach].Flags.In_Benutzung := FALSE;
       "Warenlager".Lager["HMI_Schnittstelle".Anlagendaten.Fach].Bauteil := "HMI_Schnittstelle".Anlagendaten.Bauteil;
       #tmpRD_T_ERR := RD_LOC_T("Warenlager".Lager["HMI_Schnittstelle".Anlagendaten.Fach].Zeitstempel);

       #aBeladen := FALSE;
   END_IF;
END_REGION
END_FUNCTION_BLOCK

FUNCTION_BLOCK "FC_Kran_entladen"   // FB26, FBD
{ S7_Optimized_Access := 'TRUE' }
VERSION : 0.1
   VAR_INPUT
      eKran_Ist_X : Int;
      eKran_Ist_Z : Int;
      eKran_Soll_X : Int;
      eKran_Soll_Z : Int;
      eGabel_Mitte : Bool;
      eSchrittnummer : UInt;
      ePalette_abholbereit : Bool;
   END_VAR
   VAR_OUTPUT
      aKran_Soll_X : Int;
      aKran_Soll_Z : Int;
      aGabel_Links : Bool;
      aGabel_Rechts : Bool;
      aBeladen : Bool;
   END_VAR
BEGIN

REGION Network 1 (SCL): Gabel zur Seite ausfahren
   #aGabel_Links := #eSchrittnummer = 3 OR #eSchrittnummer = 4;
END_REGION

REGION Network 2 (SCL): Gabel rechts ausfahren
   #aGabel_Rechts := #eSchrittnummer = 7 OR #eSchrittnummer = 8;
END_REGION

REGION Network 3 (SCL): Sollposition X
   // Einrichtbetrieb
   IF "HMI_Schnittstelle".Betriebsart.Einrichten THEN
       #aKran_Soll_X := "HMI_Schnittstelle".Kraene.Kran_2.Kran_Pos."X-Soll";

   // Automatikbetrieb
   ELSIF "HMI_Schnittstelle".Betriebsart.Automatik THEN

       CASE #eSchrittnummer OF
           2..5:
               //Fach mit Nummer anfahren
               #aKran_Soll_X := #eKran_Soll_X;
           ELSE:
               #aKran_Soll_X := 0;
       END_CASE;

   END_IF;
END_REGION

REGION Network 4 (SCL): Sollposition Z
   // Einrichtbetrieb
   IF "HMI_Schnittstelle".Betriebsart.Einrichten THEN
       #aKran_Soll_Z := "HMI_Schnittstelle".Kraene.Kran_2.Kran_Pos."Z-Soll";

   // Automatikbetrieb
   ELSIF "HMI_Schnittstelle".Betriebsart.Automatik THEN

       CASE #eSchrittnummer OF
           2:
               // Palette aus Fach anheben
               #aKran_Soll_Z := #eKran_Soll_Z - "Anheben_Absenken";
           4:
               //Fach mit Nummer anfahren
               #aKran_Soll_Z := #eKran_Soll_Z;
           6:
               // Palette auf Band ablegen
               #aKran_Soll_Z := "Anheben_Absenken";
           8:
               // Stapler in Grundstellung
               #aKran_Soll_Z := 0;
           ELSE:
               ;
       END_CASE;

   END_IF;
END_REGION

REGION Network 5 (SCL): Flag Kran beladen
   IF "HMI_Schnittstelle".Betriebsart.Einrichten THEN
       #"aBeladen" := FALSE;
   END_IF;


   IF #"eKran_Ist_X" = #"eKran_Soll_X"
       AND #"eKran_Ist_Z" >= #"eKran_Soll_Z" - "Anheben_Absenken"
       AND NOT #"eGabel_Mitte"
       AND NOT #"aBeladen"
   THEN
       "Warenlager".Lager["HMI_Schnittstelle".Anlagendaten.Fach].Flags.In_Benutzung := TRUE;
   END_IF;


   IF #ePalette_abholbereit
       AND #"eKran_Ist_X" = #"eKran_Soll_X"
       AND #"eKran_Ist_Z" >= #"eKran_Soll_Z"
       AND #"eGabel_Mitte"
   THEN
       #"aBeladen" := TRUE;

       "HMI_Schnittstelle".Anlagendaten.Bauteil := "Warenlager".Lager["IDB_Automatik_auslagern".Zufallszahl].Bauteil;
       "Warenlager".Lager["IDB_Automatik_auslagern".Zufallszahl] := "Warenlager".Lager[0];
   END_IF;


   IF #"eKran_Ist_X" = 0
       AND #"eKran_Ist_Z" = 0
       AND #"aBeladen"
   THEN
       "HMI_Schnittstelle".Anlagendaten.Band_aus[1] := "HMI_Schnittstelle".Anlagendaten.Bauteil;
       "HMI_Schnittstelle".Anlagendaten.Bauteil := 0;